// TIA Portal project "Pozycjoner_v7" (V15.1) (continued)
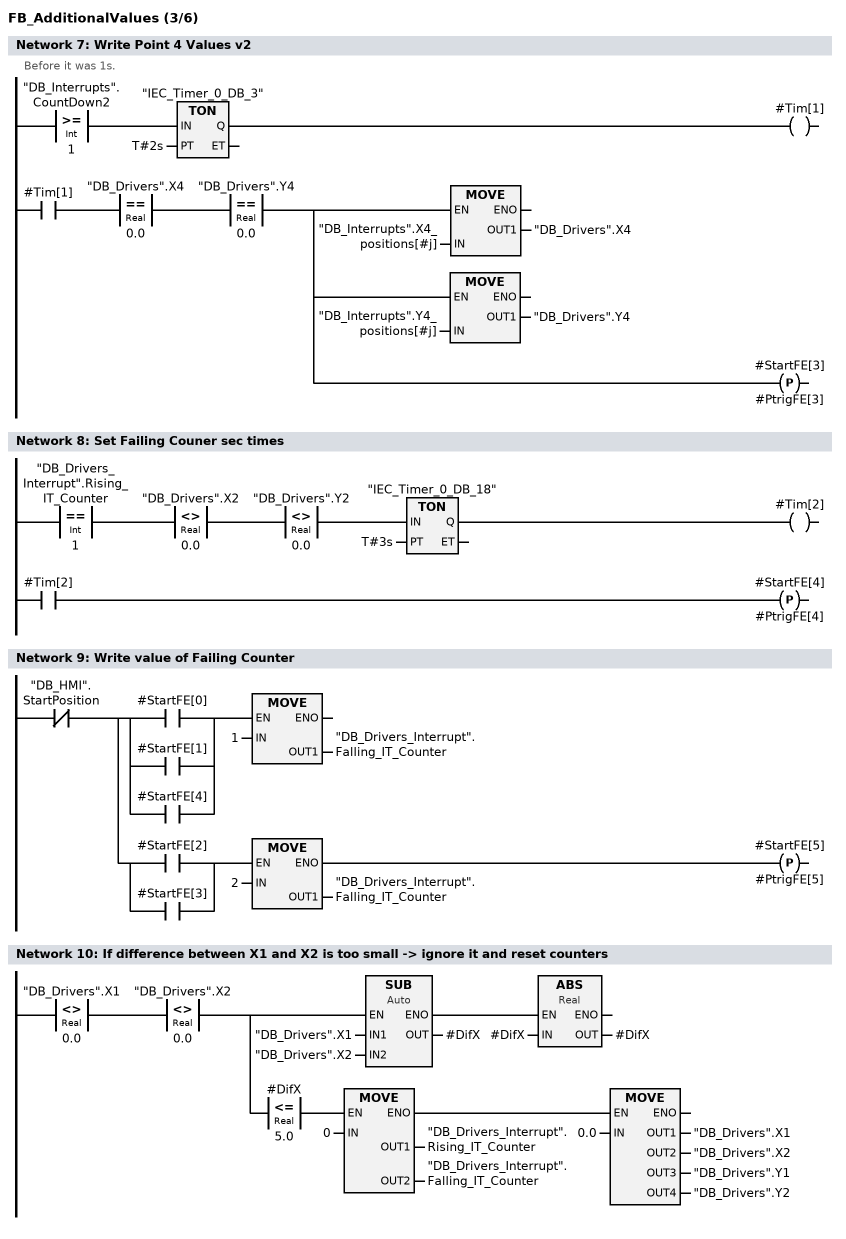
   "IEC_Timer_0_DB_3".TON(IN := "DB_Interrupts".CountDown2 >= 1, PT := T#2s);
   #Tim[1] := "IEC_Timer_0_DB_3".Q;
   #_w1 := #Tim[1] AND ("DB_Drivers".X4 = 0.0) AND ("DB_Drivers".Y4 = 0.0);
   IF #_w1 THEN
       "DB_Drivers".X4 := "DB_Interrupts".X4_positions[#j];
       "DB_Drivers".Y4 := "DB_Interrupts".Y4_positions[#j];
   END_IF;
   #StartFE[3] := #_w1 AND NOT #PtrigFE[3];   // rising edge
   #PtrigFE[3] := #_w1;
END_REGION

REGION Network 8: Set Failing Couner sec times
   "IEC_Timer_0_DB_18".TON(IN := ("DB_Drivers_Interrupt".Rising_IT_Counter = 1) AND ("DB_Drivers".X2 <> 0.0) AND ("DB_Drivers".Y2 <> 0.0),
                           PT := T#3s);
   #Tim[2] := "IEC_Timer_0_DB_18".Q;
   #StartFE[4] := #Tim[2] AND NOT #PtrigFE[4];   // rising edge
   #PtrigFE[4] := #Tim[2];
END_REGION

REGION Network 9: Write value of Failing Counter
   #_w1 := NOT "DB_HMI".StartPosition;
   IF #_w1 AND (#StartFE[0] OR #StartFE[1] OR #StartFE[4]) THEN
       "DB_Drivers_Interrupt".Falling_IT_Counter := 1;
   END_IF;
   #_w2 := #_w1 AND (#StartFE[2] OR #StartFE[3]);
   IF #_w2 THEN "DB_Drivers_Interrupt".Falling_IT_Counter := 2; END_IF;
   #StartFE[5] := #_w2 AND NOT #PtrigFE[5];   // rising edge
   #PtrigFE[5] := #_w2;
END_REGION

REGION Network 10: If difference between X1 and X2 is too small -> ignore it and reset counters
   RUNG wire#powerrail
      { S7_Templates := "SrcType := Real" } NE_Contact(in1 := "DB_Drivers".X1, in2 := 0.0)
      { S7_Templates := "SrcType := Real" } NE_Contact(in1 := "DB_Drivers".X2, in2 := 0.0)
      wire#w1
      Sub(in1 := "DB_Drivers".X1, in2 := "DB_Drivers".X2, out => #DifX)
      { S7_Templates := "SrcType := Real" } Abs(in := #DifX, out => #DifX)
   END_RUNG
   RUNG wire#w1
      { S7_Templates := "SrcType := Real" } LE_Contact(in1 := #DifX, in2 := 5.0)
      Move(in := 0, out1 => "DB_Drivers_Interrupt".Rising_IT_Counter, out2 => "DB_Drivers_Interrupt".Falling_IT_Counter)
      Move(in := 0.0, out1 => "DB_Drivers".X1, out2 => "DB_Drivers".X2, out3 => "DB_Drivers".Y1, out4 => "DB_Drivers".Y2)
   END_RUNG
   // the same network as SCL:
   #_w1 := ("DB_Drivers".X1 <> 0.0) AND ("DB_Drivers".X2 <> 0.0);
   IF #_w1 THEN
       #DifX := "DB_Drivers".X1 - "DB_Drivers".X2;
       #DifX := ABS(#DifX);
   END_IF;
   IF #_w1 AND (#DifX <= 5.0) THEN
       "DB_Drivers_Interrupt".Rising_IT_Counter := 0;
       "DB_Drivers_Interrupt".Falling_IT_Counter := 0;
       "DB_Drivers".X1 := 0.0;
       "DB_Drivers".X2 := 0.0;
       "DB_Drivers".Y1 := 0.0;
       "DB_Drivers".Y2 := 0.0;
   END_IF;
END_REGION

REGION Network 11: Repeat move if rising edge was detected but falling edge counter = 0 for 10 sec
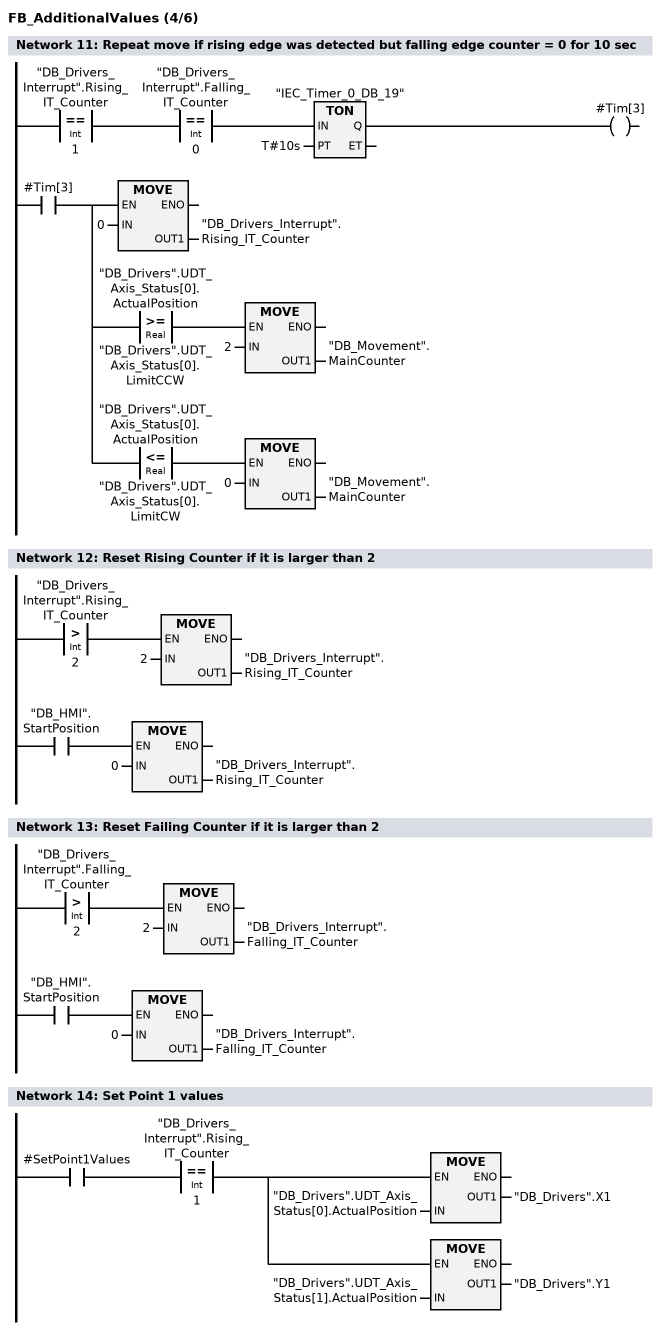
   "IEC_Timer_0_DB_19".TON(IN := ("DB_Drivers_Interrupt".Rising_IT_Counter = 1) AND ("DB_Drivers_Interrupt".Falling_IT_Counter = 0),
                           PT := T#10s);
   #Tim[3] := "IEC_Timer_0_DB_19".Q;
   IF #Tim[3] THEN "DB_Drivers_Interrupt".Rising_IT_Counter := 0; END_IF;
   IF #Tim[3] AND ("DB_Drivers".UDT_Axis_Status[0].ActualPosition >= "DB_Drivers".UDT_Axis_Status[0].LimitCCW) THEN
       "DB_Movement".MainCounter := 2;
   END_IF;
   IF #Tim[3] AND ("DB_Drivers".UDT_Axis_Status[0].ActualPosition <= "DB_Drivers".UDT_Axis_Status[0].LimitCW) THEN
       "DB_Movement".MainCounter := 0;
   END_IF;
END_REGION

REGION Network 12: Reset Rising Counter if it is larger than 2
   RUNG wire#powerrail
      { S7_Templates := "SrcType := Int" } GT_Contact(in1 := "DB_Drivers_Interrupt".Rising_IT_Counter, in2 := 2)
      Move(in := 2, out1 => "DB_Drivers_Interrupt".Rising_IT_Counter)
   END_RUNG
   RUNG wire#powerrail
      Contact( "DB_HMI".StartPosition )
      Move(in := 0, out1 => "DB_Drivers_Interrupt".Rising_IT_Counter)
   END_RUNG
   // the same network as SCL:
   IF "DB_Drivers_Interrupt".Rising_IT_Counter > 2 THEN
       "DB_Drivers_Interrupt".Rising_IT_Counter := 2;
   END_IF;
   IF "DB_HMI".StartPosition THEN "DB_Drivers_Interrupt".Rising_IT_Counter := 0; END_IF;
END_REGION

REGION Network 13: Reset Failing Counter if it is larger than 2
   RUNG wire#powerrail
      { S7_Templates := "SrcType := Int" } GT_Contact(in1 := "DB_Drivers_Interrupt".Falling_IT_Counter, in2 := 2)
      Move(in := 2, out1 => "DB_Drivers_Interrupt".Falling_IT_Counter)
   END_RUNG
   RUNG wire#powerrail
      Contact( "DB_HMI".StartPosition )
      Move(in := 0, out1 => "DB_Drivers_Interrupt".Falling_IT_Counter)
   END_RUNG
   // the same network as SCL:
   IF "DB_Drivers_Interrupt".Falling_IT_Counter > 2 THEN
       "DB_Drivers_Interrupt".Falling_IT_Counter := 2;
   END_IF;
   IF "DB_HMI".StartPosition THEN "DB_Drivers_Interrupt".Falling_IT_Counter := 0; END_IF;
END_REGION

REGION Network 14: Set Point 1 values
   RUNG wire#powerrail
      Contact( #SetPoint1Values )
      { S7_Templates := "SrcType := Int" } EQ_Contact(in1 := "DB_Drivers_Interrupt".Rising_IT_Counter, in2 := 1)
      wire#w1
      Move(in := "DB_Drivers".UDT_Axis_Status[0].ActualPosition, out1 => "DB_Drivers".X1)
   END_RUNG
   RUNG wire#w1
      Move(in := "DB_Drivers".UDT_Axis_Status[1].ActualPosition, out1 => "DB_Drivers".Y1)
   END_RUNG
   // the same network as SCL:
   IF #SetPoint1Values AND ("DB_Drivers_Interrupt".Rising_IT_Counter = 1) THEN
       "DB_Drivers".X1 := "DB_Drivers".UDT_Axis_Status[0].ActualPosition;
       "DB_Drivers".Y1 := "DB_Drivers".UDT_Axis_Status[1].ActualPosition;
   END_IF;
END_REGION

REGION Network 15: Set Point 3 values
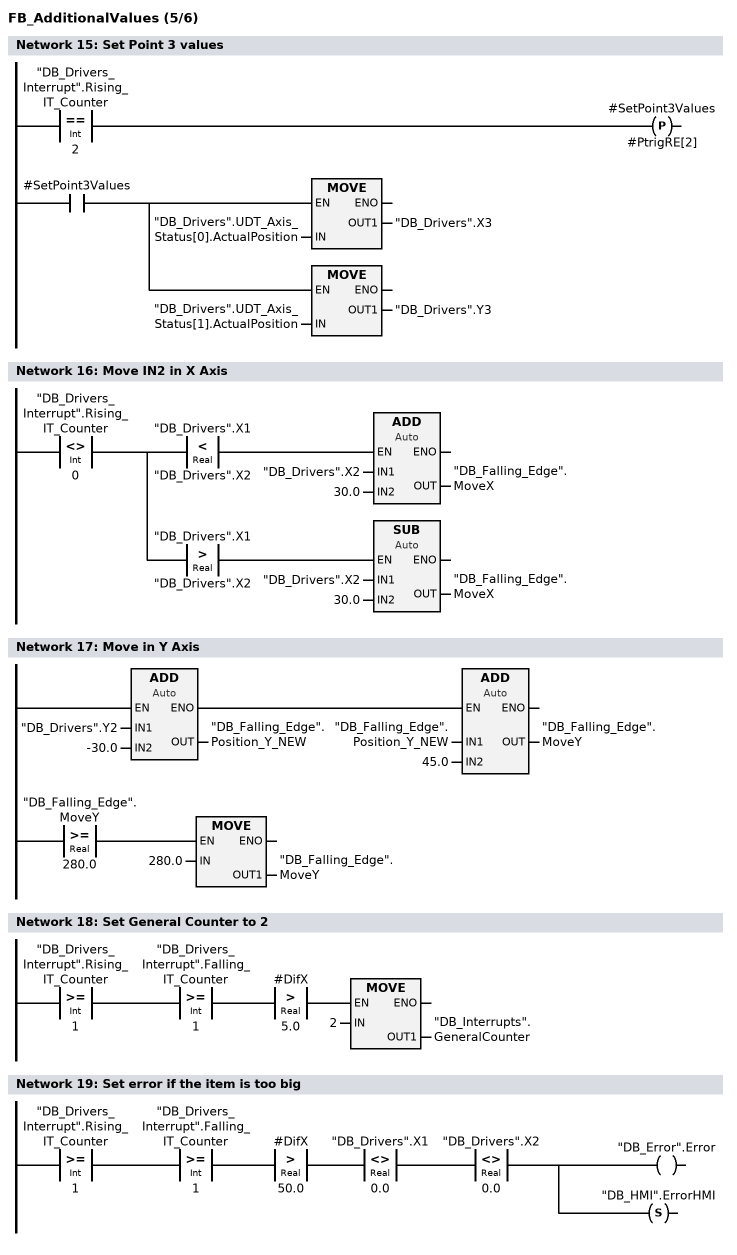
   #_w1 := "DB_Drivers_Interrupt".Rising_IT_Counter = 2;
   #SetPoint3Values := #_w1 AND NOT #PtrigRE[2];   // rising edge
   #PtrigRE[2] := #_w1;
   IF #SetPoint3Values THEN
       "DB_Drivers".X3 := "DB_Drivers".UDT_Axis_Status[0].ActualPosition;
       "DB_Drivers".Y3 := "DB_Drivers".UDT_Axis_Status[1].ActualPosition;
   END_IF;
END_REGION

REGION Network 16: Move IN2 in X Axis
   RUNG wire#powerrail
      { S7_Templates := "SrcType := Int" } NE_Contact(in1 := "DB_Drivers_Interrupt".Rising_IT_Counter, in2 := 0)
      wire#w1
      { S7_Templates := "SrcType := Real" } LT_Contact(in1 := "DB_Drivers".X1, in2 := "DB_Drivers".X2)
      Add(in1 := "DB_Drivers".X2, in2 := 30.0, out => "DB_Falling_Edge".MoveX)
   END_RUNG
   RUNG wire#w1
      { S7_Templates := "SrcType := Real" } GT_Contact(in1 := "DB_Drivers".X1, in2 := "DB_Drivers".X2)
      Sub(in1 := "DB_Drivers".X2, in2 := 30.0, out => "DB_Falling_Edge".MoveX)
   END_RUNG
   // the same network as SCL:
   #_w1 := "DB_Drivers_Interrupt".Rising_IT_Counter <> 0;
   IF #_w1 AND ("DB_Drivers".X1 < "DB_Drivers".X2) THEN
       "DB_Falling_Edge".MoveX := "DB_Drivers".X2 + 30.0;
   END_IF;
   IF #_w1 AND ("DB_Drivers".X1 > "DB_Drivers".X2) THEN
       "DB_Falling_Edge".MoveX := "DB_Drivers".X2 - 30.0;
   END_IF;
END_REGION

REGION Network 17: Move in Y Axis
   RUNG wire#powerrail
      Add(in1 := "DB_Drivers".Y2, in2 := -30.0, out => "DB_Falling_Edge".Position_Y_NEW)
      Add(in1 := "DB_Falling_Edge".Position_Y_NEW, in2 := 45.0, out => "DB_Falling_Edge".MoveY)
   END_RUNG
   RUNG wire#powerrail
      { S7_Templates := "SrcType := Real" } GE_Contact(in1 := "DB_Falling_Edge".MoveY, in2 := 280.0)
      Move(in := 280.0, out1 => "DB_Falling_Edge".MoveY)
   END_RUNG
   // the same network as SCL:
   "DB_Falling_Edge".Position_Y_NEW := "DB_Drivers".Y2 + (-30.0);
   "DB_Falling_Edge".MoveY := "DB_Falling_Edge".Position_Y_NEW + 45.0;
   IF "DB_Falling_Edge".MoveY >= 280.0 THEN "DB_Falling_Edge".MoveY := 280.0; END_IF;
END_REGION

REGION Network 18: Set General Counter to 2
   RUNG wire#powerrail
      { S7_Templates := "SrcType := Int" } GE_Contact(in1 := "DB_Drivers_Interrupt".Rising_IT_Counter, in2 := 1)
      { S7_Templates := "SrcType := Int" } GE_Contact(in1 := "DB_Drivers_Interrupt".Falling_IT_Counter, in2 := 1)
      { S7_Templates := "SrcType := Real" } GT_Contact(in1 := #DifX, in2 := 5.0)
      Move(in := 2, out1 => "DB_Interrupts".GeneralCounter)
   END_RUNG
   // the same network as SCL:
   IF ("DB_Drivers_Interrupt".Rising_IT_Counter >= 1) AND ("DB_Drivers_Interrupt".Falling_IT_Counter >= 1) AND (#DifX > 5.0) THEN
       "DB_Interrupts".GeneralCounter := 2;
   END_IF;
END_REGION

REGION Network 19: Set error if the item is too big
   RUNG wire#powerrail
      { S7_Templates := "SrcType := Int" } GE_Contact(in1 := "DB_Drivers_Interrupt".Rising_IT_Counter, in2 := 1)
      { S7_Templates := "SrcType := Int" } GE_Contact(in1 := "DB_Drivers_Interrupt".Falling_IT_Counter, in2 := 1)
      { S7_Templates := "SrcType := Real" } GT_Contact(in1 := #DifX, in2 := 50.0)
      { S7_Templates := "SrcType := Real" } NE_Contact(in1 := "DB_Drivers".X1, in2 := 0.0)
      { S7_Templates := "SrcType := Real" } NE_Contact(in1 := "DB_Drivers".X2, in2 := 0.0)
      wire#w1
      Coil( "DB_Error".Error )
   END_RUNG
   RUNG wire#w1
      S_Coil( "DB_HMI".ErrorHMI )
   END_RUNG
   // the same network as SCL:
   "DB_Error".Error := ("DB_Drivers_Interrupt".Rising_IT_Counter >= 1) AND ("DB_Drivers_Interrupt".Falling_IT_Counter >= 1) AND (#DifX > 50.0) AND ("DB_Drivers".X1 <> 0.0) AND ("DB_Drivers".X2 <> 0.0);
   IF "DB_Error".Error THEN "DB_HMI".ErrorHMI := TRUE; END_IF;
END_REGION

REGION Network 20: Check the last point once again
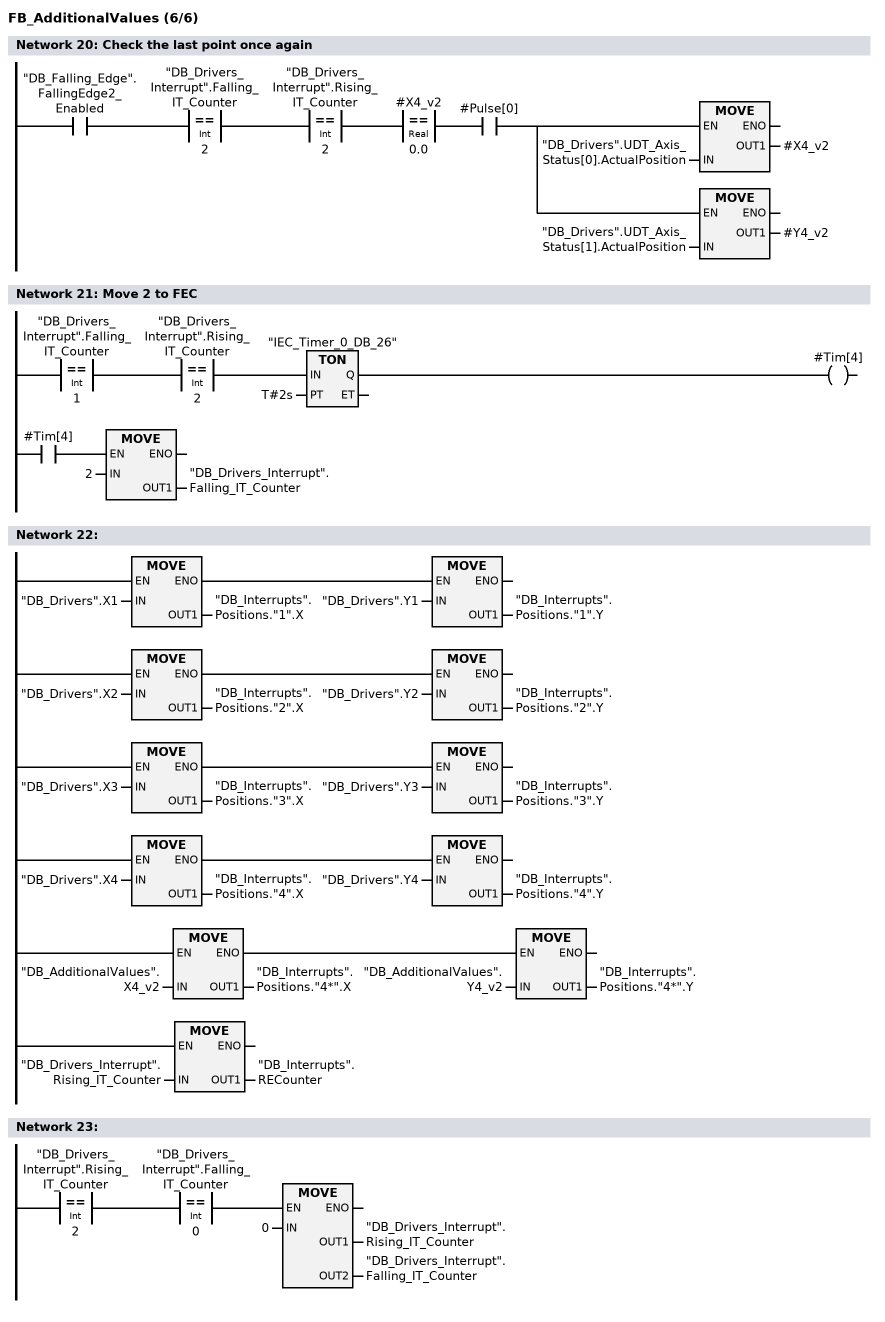
   RUNG wire#powerrail
      Contact( "DB_Falling_Edge".FallingEdge2_Enabled )
      { S7_Templates := "SrcType := Int" } EQ_Contact(in1 := "DB_Drivers_Interrupt".Falling_IT_Counter, in2 := 2)
      { S7_Templates := "SrcType := Int" } EQ_Contact(in1 := "DB_Drivers_Interrupt".Rising_IT_Counter, in2 := 2)
      { S7_Templates := "SrcType := Real" } EQ_Contact(in1 := #X4_v2, in2 := 0.0)
      Contact( #Pulse[0] )
      wire#w1
      Move(in := "DB_Drivers".UDT_Axis_Status[0].ActualPosition, out1 => #X4_v2)
   END_RUNG
   RUNG wire#w1
      Move(in := "DB_Drivers".UDT_Axis_Status[1].ActualPosition, out1 => #Y4_v2)
   END_RUNG
   // the same network as SCL:
   #_w1 := "DB_Falling_Edge".FallingEdge2_Enabled AND ("DB_Drivers_Interrupt".Falling_IT_Counter = 2) AND ("DB_Drivers_Interrupt".Rising_IT_Counter = 2) AND (#X4_v2 = 0.0) AND #Pulse[0];
   IF #_w1 THEN
       #X4_v2 := "DB_Drivers".UDT_Axis_Status[0].ActualPosition;
       #Y4_v2 := "DB_Drivers".UDT_Axis_Status[1].ActualPosition;
   END_IF;
END_REGION

REGION Network 21: Move 2 to FEC
   "IEC_Timer_0_DB_26".TON(IN := ("DB_Drivers_Interrupt".Falling_IT_Counter = 1) AND ("DB_Drivers_Interrupt".Rising_IT_Counter = 2),
                           PT := T#2s);
   #Tim[4] := "IEC_Timer_0_DB_26".Q;
   IF #Tim[4] THEN "DB_Drivers_Interrupt".Falling_IT_Counter := 2; END_IF;
END_REGION

REGION Network 22
   RUNG wire#powerrail
      Move(in := "DB_Drivers".X1, out1 => "DB_Interrupts".Positions."1".X)
      Move(in := "DB_Drivers".Y1, out1 => "DB_Interrupts".Positions."1".Y)
   END_RUNG
   RUNG wire#powerrail
      Move(in := "DB_Drivers".X2, out1 => "DB_Interrupts".Positions."2".X)
      Move(in := "DB_Drivers".Y2, out1 => "DB_Interrupts".Positions."2".Y)
   END_RUNG
   RUNG wire#powerrail
      Move(in := "DB_Drivers".X3, out1 => "DB_Interrupts".Positions."3".X)
      Move(in := "DB_Drivers".Y3, out1 => "DB_Interrupts".Positions."3".Y)
   END_RUNG
   RUNG wire#powerrail
      Move(in := "DB_Drivers".X4, out1 => "DB_Interrupts".Positions."4".X)
      Move(in := "DB_Drivers".Y4, out1 => "DB_Interrupts".Positions."4".Y)
   END_RUNG
   RUNG wire#powerrail
      Move(in := "DB_AdditionalValues".X4_v2, out1 => "DB_Interrupts".Positions."4*".X)
      Move(in := "DB_AdditionalValues".Y4_v2, out1 => "DB_Interrupts".Positions."4*".Y)
   END_RUNG
   RUNG wire#powerrail
      Move(in := "DB_Drivers_Interrupt".Rising_IT_Counter, out1 => "DB_Interrupts".RECounter)
   END_RUNG
   // the same network as SCL:
   "DB_Interrupts".Positions."1".X := "DB_Drivers".X1;
   "DB_Interrupts".Positions."1".Y := "DB_Drivers".Y1;
   "DB_Interrupts".Positions."2".X := "DB_Drivers".X2;
   "DB_Interrupts".Positions."2".Y := "DB_Drivers".Y2;
   "DB_Interrupts".Positions."3".X := "DB_Drivers".X3;
   "DB_Interrupts".Positions."3".Y := "DB_Drivers".Y3;
   "DB_Interrupts".Positions."4".X := "DB_Drivers".X4;
   "DB_Interrupts".Positions."4".Y := "DB_Drivers".Y4;
   "DB_Interrupts".Positions."4*".X := "DB_AdditionalValues".X4_v2;
   "DB_Interrupts".Positions."4*".Y := "DB_AdditionalValues".Y4_v2;
   "DB_Interrupts".RECounter := "DB_Drivers_Interrupt".Rising_IT_Counter;
END_REGION

REGION Network 23
   RUNG wire#powerrail
      { S7_Templates := "SrcType := Int" } EQ_Contact(in1 := "DB_Drivers_Interrupt".Rising_IT_Counter, in2 := 2)
      { S7_Templates := "SrcType := Int" } EQ_Contact(in1 := "DB_Drivers_Interrupt".Falling_IT_Counter, in2 := 0)
      Move(in := 0, out1 => "DB_Drivers_Interrupt".Rising_IT_Counter, out2 => "DB_Drivers_Interrupt".Falling_IT_Counter)
   END_RUNG
   // the same network as SCL:
   IF ("DB_Drivers_Interrupt".Rising_IT_Counter = 2) AND ("DB_Drivers_Interrupt".Falling_IT_Counter = 0) THEN
       "DB_Drivers_Interrupt".Rising_IT_Counter := 0;
       "DB_Drivers_Interrupt".Falling_IT_Counter := 0;
   END_IF;
END_REGION
END_FUNCTION_BLOCK

FUNCTION_BLOCK "FB_Falling_Edge"   // FB9, LAD
{ S7_Optimized_Access := 'TRUE' }
VERSION : 0.1
   VAR_INPUT
      LaserSensor : Bool;
   END_VAR
   VAR
      X_Position2 : Real;
      Y_Position2 : Real;
      Position_Y_NEW : Real;   // New Y position
      MoveX : Real;   // Keep moving after detecting item
      UDT_AxisControl : Array[0..2] of "UDT_AxisControl";
      UDT_AxisStatus : Array[0..2] of "UDT_AxisStatus";
      Y_MIN : Int;
      Y_MAX : Real;
      MoveX_MIN : Int;
      MoveX_MAX : Int;
      MoveY : Real;
      MainCounter : Int;
      Enabled : Bool;
      moveY_min : Int;
      moveY_max : Int;
      FallingEdge2_Enabled : Bool;
      StartX : Array[0..2] of Bool;
      StartY : Array[0..2] of Bool;
      PtrigX : Array[0..2] of Bool;
      PtrigY : Array[0..2] of Bool;
      Timers : Array[0..2] of Bool;
   END_VAR
   VAR_TEMP   // added for the SCL form of the ladder/FBD networks
      _w1 : Bool;
   END_VAR
BEGIN

REGION Network 1: Enabled
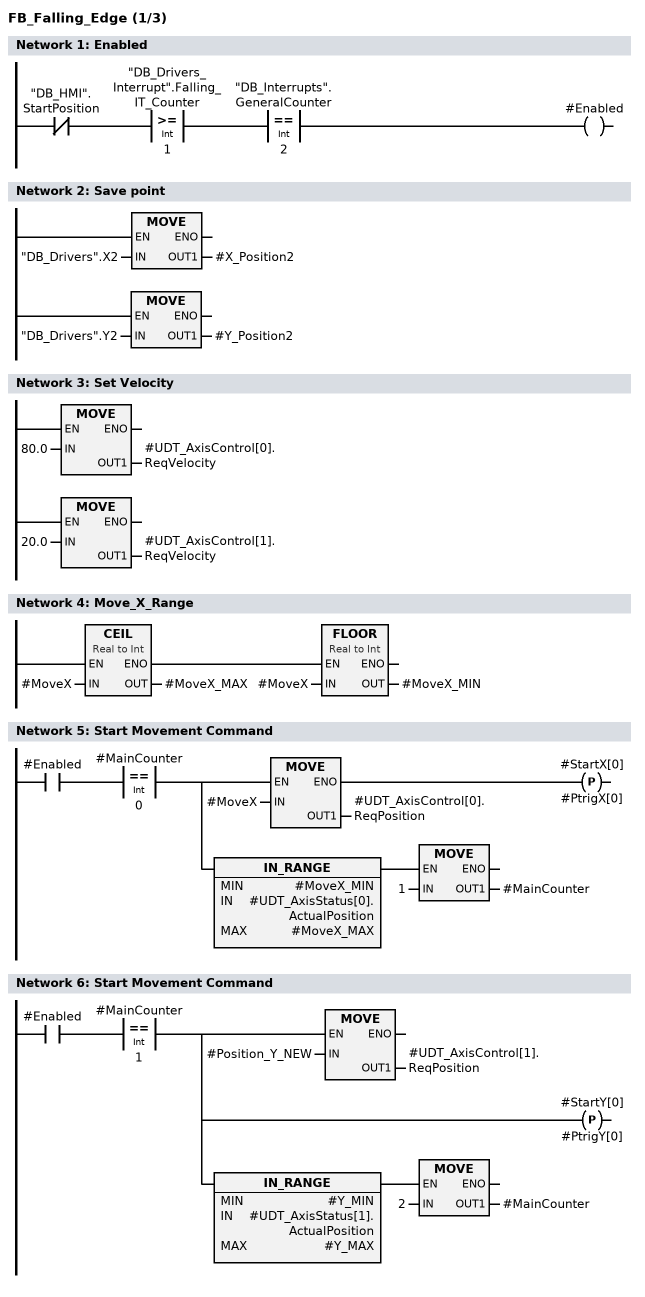
   RUNG wire#powerrail
      I_Contact( "DB_HMI".StartPosition )
      { S7_Templates := "SrcType := Int" } GE_Contact(in1 := "DB_Drivers_Interrupt".Falling_IT_Counter, in2 := 1)
      { S7_Templates := "SrcType := Int" } EQ_Contact(in1 := "DB_Interrupts".GeneralCounter, in2 := 2)
      Coil( #Enabled )
   END_RUNG
   // the same network as SCL:
   #Enabled := NOT "DB_HMI".StartPosition AND ("DB_Drivers_Interrupt".Falling_IT_Counter >= 1) AND ("DB_Interrupts".GeneralCounter = 2);
END_REGION

REGION Network 2: Save point
   RUNG wire#powerrail
      Move(in := "DB_Drivers".X2, out1 => #X_Position2)
   END_RUNG
   RUNG wire#powerrail
      Move(in := "DB_Drivers".Y2, out1 => #Y_Position2)
   END_RUNG
   // the same network as SCL:
   #X_Position2 := "DB_Drivers".X2;
   #Y_Position2 := "DB_Drivers".Y2;
END_REGION

REGION Network 3: Set Velocity
   RUNG wire#powerrail
      Move(in := 80.0, out1 => #UDT_AxisControl[0].ReqVelocity)
   END_RUNG
   RUNG wire#powerrail
      Move(in := 20.0, out1 => #UDT_AxisControl[1].ReqVelocity)
   END_RUNG
   // the same network as SCL:
   #UDT_AxisControl[0].ReqVelocity := 80.0;
   #UDT_AxisControl[1].ReqVelocity := 20.0;
END_REGION

REGION Network 4: Move_X_Range
   #MoveX_MAX := CEIL(#MoveX);
   #MoveX_MIN := FLOOR(#MoveX);
END_REGION

REGION Network 5: Start Movement Command
   #_w1 := #Enabled AND (#MainCounter = 0);
   IF #_w1 THEN #UDT_AxisControl[0].ReqPosition := #MoveX; END_IF;
   #StartX[0] := #_w1 AND NOT #PtrigX[0];   // rising edge
   #PtrigX[0] := #_w1;
   IF #_w1 AND (#MoveX_MIN <= #UDT_AxisStatus[0].ActualPosition) AND (#UDT_AxisStatus[0].ActualPosition <= #MoveX_MAX) THEN
       #MainCounter := 1;
   END_IF;
END_REGION

REGION Network 6: Start Movement Command
   #_w1 := #Enabled AND (#MainCounter = 1);
   IF #_w1 THEN #UDT_AxisControl[1].ReqPosition := #Position_Y_NEW; END_IF;
   #StartY[0] := #_w1 AND NOT #PtrigY[0];   // rising edge
   #PtrigY[0] := #_w1;
   IF #_w1 AND (#Y_MIN <= #UDT_AxisStatus[1].ActualPosition) AND (#UDT_AxisStatus[1].ActualPosition <= #Y_MAX) THEN
       #MainCounter := 2;
   END_IF;
END_REGION

REGION Network 7: NewPositionY Range
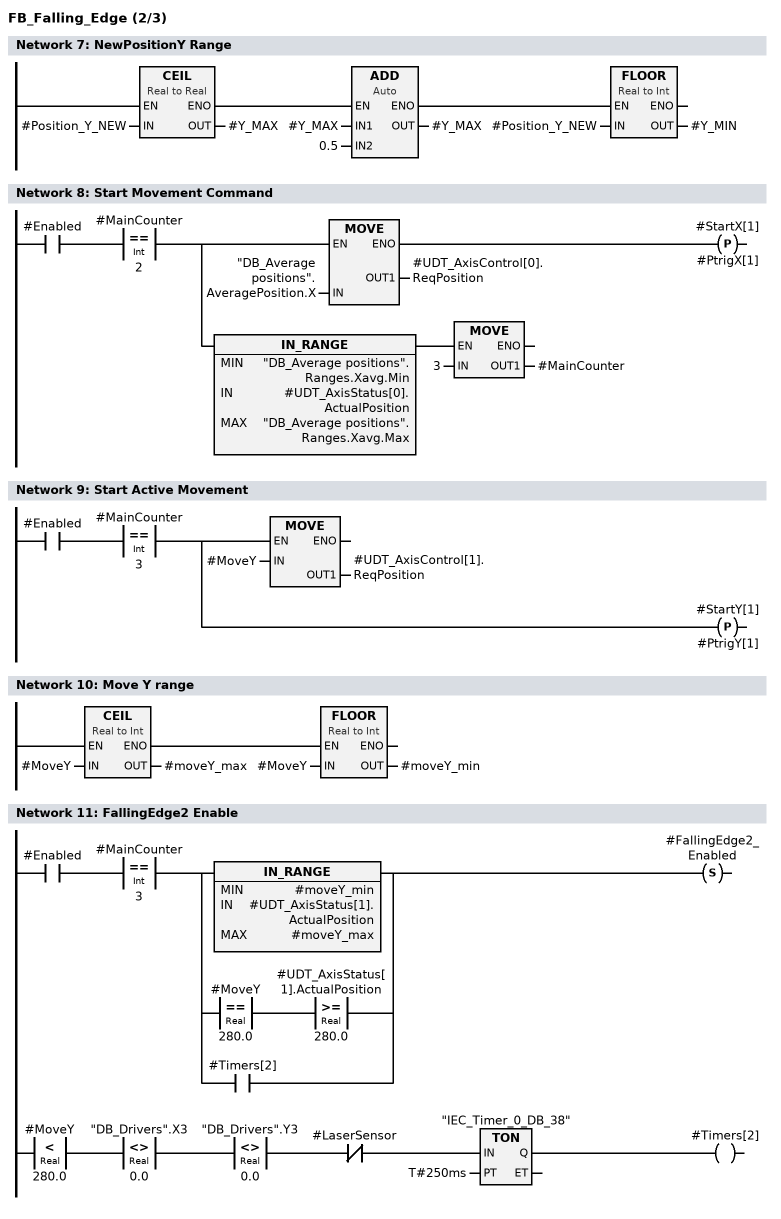
   #Y_MAX := CEIL(#Position_Y_NEW);
   #Y_MAX := #Y_MAX + 0.5;
   #Y_MIN := FLOOR(#Position_Y_NEW);
END_REGION

REGION Network 8: Start Movement Command
   #_w1 := #Enabled AND (#MainCounter = 2);
   IF #_w1 THEN #UDT_AxisControl[0].ReqPosition := "DB_Average positions".AveragePosition.X; END_IF;
   #StartX[1] := #_w1 AND NOT #PtrigX[1];   // rising edge
   #PtrigX[1] := #_w1;
   IF #_w1 AND ("DB_Average positions".Ranges.Xavg.Min <= #UDT_AxisStatus[0].ActualPosition) AND (#UDT_AxisStatus[0].ActualPosition <= "DB_Average positions".Ranges.Xavg.Max) THEN
       #MainCounter := 3;
   END_IF;
END_REGION

REGION Network 9: Start Active Movement
   #_w1 := #Enabled AND (#MainCounter = 3);
   IF #_w1 THEN #UDT_AxisControl[1].ReqPosition := #MoveY; END_IF;
   #StartY[1] := #_w1 AND NOT #PtrigY[1];   // rising edge
   #PtrigY[1] := #_w1;
END_REGION

REGION Network 10: Move Y range
   #moveY_max := CEIL(#MoveY);
   #moveY_min := FLOOR(#MoveY);
END_REGION

REGION Network 11: FallingEdge2 Enable
   IF #Enabled AND (#MainCounter = 3) AND (((#moveY_min <= #UDT_AxisStatus[1].ActualPosition) AND (#UDT_AxisStatus[1].ActualPosition <= #moveY_max)) OR ((#MoveY = 280.0) AND (#UDT_AxisStatus[1].ActualPosition >= 280.0)) OR #Timers[2]) THEN
       #FallingEdge2_Enabled := TRUE;
   END_IF;
   "IEC_Timer_0_DB_38".TON(IN := (#MoveY < 280.0) AND ("DB_Drivers".X3 <> 0.0) AND ("DB_Drivers".Y3 <> 0.0) AND NOT #LaserSensor,
                           PT := T#250ms);
   #Timers[2] := "IEC_Timer_0_DB_38".Q;
END_REGION

REGION Network 12: Start Movement Command
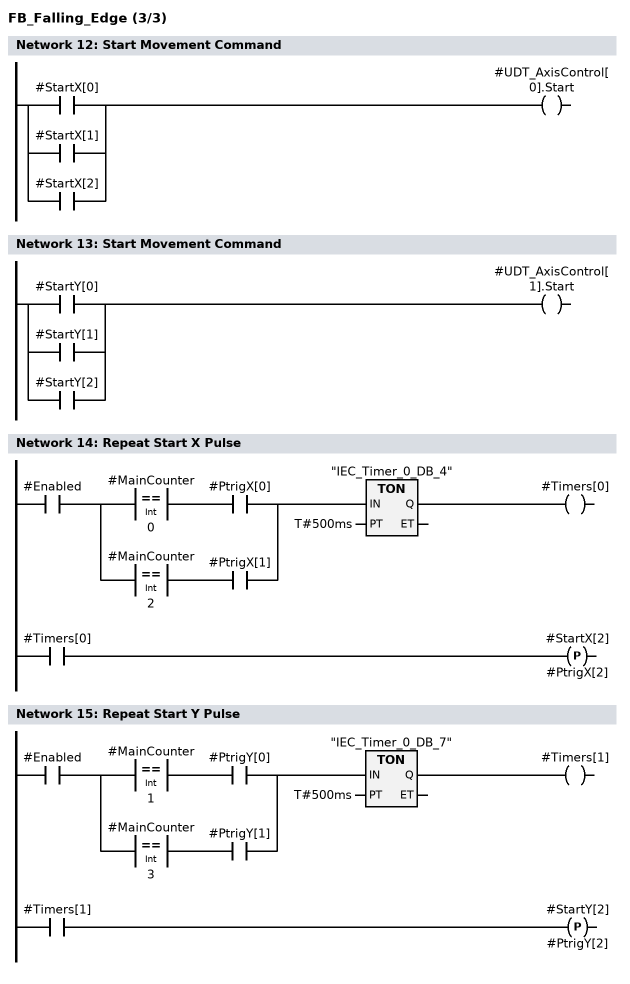
   RUNG wire#powerrail
      Contact( #StartX[0] )
      wire#w1
      Coil( #UDT_AxisControl[0].Start )
   END_RUNG
   RUNG wire#powerrail
      Contact( #StartX[1] )
   END_RUNG wire#w1
   RUNG wire#powerrail
      Contact( #StartX[2] )
   END_RUNG wire#w1
   // the same network as SCL:
   #UDT_AxisControl[0].Start := #StartX[0] OR #StartX[1] OR #StartX[2];
END_REGION

REGION Network 13: Start Movement Command
   RUNG wire#powerrail
      Contact( #StartY[0] )
      wire#w1
      Coil( #UDT_AxisControl[1].Start )
   END_RUNG
   RUNG wire#powerrail
      Contact( #StartY[1] )
   END_RUNG wire#w1
   RUNG wire#powerrail
      Contact( #StartY[2] )
   END_RUNG wire#w1
   // the same network as SCL:
   #UDT_AxisControl[1].Start := #StartY[0] OR #StartY[1] OR #StartY[2];
END_REGION

REGION Network 14: Repeat Start X Pulse
   "IEC_Timer_0_DB_4".TON(IN := #Enabled AND (((#MainCounter = 0) AND #PtrigX[0]) OR ((#MainCounter = 2) AND #PtrigX[1])),
                          PT := T#500ms);
   #Timers[0] := "IEC_Timer_0_DB_4".Q;
   #StartX[2] := #Timers[0] AND NOT #PtrigX[2];   // rising edge
   #PtrigX[2] := #Timers[0];
END_REGION

REGION Network 15: Repeat Start Y Pulse
   "IEC_Timer_0_DB_7".TON(IN := #Enabled AND (((#MainCounter = 1) AND #PtrigY[0]) OR ((#MainCounter = 3) AND #PtrigY[1])),
                          PT := T#500ms);
   #Timers[1] := "IEC_Timer_0_DB_7".Q;
   #StartY[2] := #Timers[1] AND NOT #PtrigY[2];   // rising edge
   #PtrigY[2] := #Timers[1];
END_REGION
END_FUNCTION_BLOCK

// folder: Displacement/Center Point Calculation/Line2

FUNCTION_BLOCK "FB_Line2"   // FB11, LAD
{ S7_Optimized_Access := 'TRUE' }
VERSION : 0.1
   VAR_INPUT
      LaserSensor : Bool;
   END_VAR
   VAR
      UDT_AxisControl : Array[0..2] of "UDT_AxisControl";
      UDT_AxisStatus : Array[0..2] of "UDT_AxisStatus";
      Ranges : Struct
         X_MAX : Real;
         X_MIN : Real;
         Y_MAX : Real;
         Y_MIN : Real;
      END_STRUCT;
      StartX : Array[0..3] of Bool;
      PtrigX : Array[0..3] of Bool;
      StartY : Array[0..4] of Bool;
      PtrigY : Array[0..4] of Bool;
      Enabled : Bool;
      Midpoint : Bool;
      Tim : Array[0..5] of Bool;
   END_VAR
   VAR_TEMP   // added for the SCL form of the ladder/FBD networks
      _w1 : Bool;
      _w2 : Bool;
   END_VAR
BEGIN

REGION Network 1: Enabled block
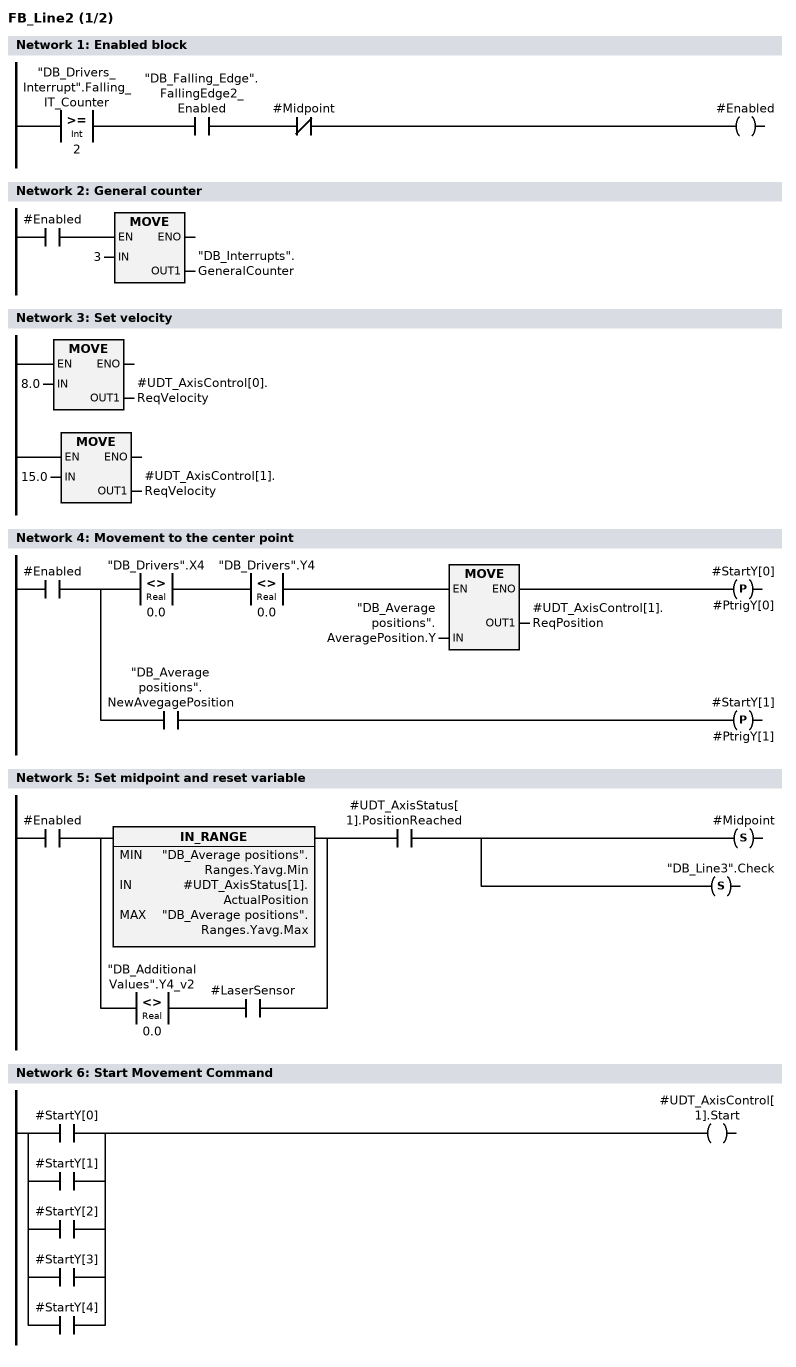
   RUNG wire#powerrail
      { S7_Templates := "SrcType := Int" } GE_Contact(in1 := "DB_Drivers_Interrupt".Falling_IT_Counter, in2 := 2)
      Contact( "DB_Falling_Edge".FallingEdge2_Enabled )
      I_Contact( #Midpoint )
      Coil( #Enabled )
   END_RUNG
   // the same network as SCL:
   #Enabled := ("DB_Drivers_Interrupt".Falling_IT_Counter >= 2) AND "DB_Falling_Edge".FallingEdge2_Enabled AND NOT #Midpoint;
END_REGION

REGION Network 2: General counter
   RUNG wire#powerrail
      Contact( #Enabled )
      Move(in := 3, out1 => "DB_Interrupts".GeneralCounter)
   END_RUNG
   // the same network as SCL:
   IF #Enabled THEN "DB_Interrupts".GeneralCounter := 3; END_IF;
END_REGION

REGION Network 3: Set velocity
   RUNG wire#powerrail
      Move(in := 8.0, out1 => #UDT_AxisControl[0].ReqVelocity)
   END_RUNG
   RUNG wire#powerrail
      Move(in := 15.0, out1 => #UDT_AxisControl[1].ReqVelocity)
   END_RUNG
   // the same network as SCL:
   #UDT_AxisControl[0].ReqVelocity := 8.0;
   #UDT_AxisControl[1].ReqVelocity := 15.0;
END_REGION

REGION Network 4: Movement to the center point
   #_w1 := #Enabled AND ("DB_Drivers".X4 <> 0.0) AND ("DB_Drivers".Y4 <> 0.0);
   IF #_w1 THEN #UDT_AxisControl[1].ReqPosition := "DB_Average positions".AveragePosition.Y; END_IF;
   #StartY[0] := #_w1 AND NOT #PtrigY[0];   // rising edge
   #PtrigY[0] := #_w1;
   #_w2 := #Enabled AND "DB_Average positions".NewAvegagePosition;
   #StartY[1] := #_w2 AND NOT #PtrigY[1];   // rising edge
   #PtrigY[1] := #_w2;
END_REGION

REGION Network 5: Set midpoint and reset variable
   RUNG wire#powerrail
      Contact( #Enabled )
      wire#w1
      { S7_Templates := "SrcType := Real" } InRange(min := "DB_Average positions".Ranges.Yavg.Min, in := #UDT_AxisStatus[1].ActualPosition, max := "DB_Average positions".Ranges.Yavg.Max)
      wire#w2
      Contact( #UDT_AxisStatus[1].PositionReached )
      wire#w3
      S_Coil( #Midpoint )
   END_RUNG
   RUNG wire#w1
      { S7_Templates := "SrcType := Real" } NE_Contact(in1 := "DB_AdditionalValues".Y4_v2, in2 := 0.0)
      Contact( #LaserSensor )
   END_RUNG wire#w2
   RUNG wire#w3
      S_Coil( "DB_Line3".Check )
   END_RUNG
   // the same network as SCL:
   IF #Enabled AND ((("DB_Average positions".Ranges.Yavg.Min <= #UDT_AxisStatus[1].ActualPosition) AND (#UDT_AxisStatus[1].ActualPosition <= "DB_Average positions".Ranges.Yavg.Max)) OR (("DB_AdditionalValues".Y4_v2 <> 0.0) AND #LaserSensor)) AND #UDT_AxisStatus[1].PositionReached THEN
       #Midpoint := TRUE;
       "DB_Line3".Check := TRUE;
   END_IF;
END_REGION

REGION Network 6: Start Movement Command
   RUNG wire#powerrail
      Contact( #StartY[0] )
      wire#w1
      Coil( #UDT_AxisControl[1].Start )
   END_RUNG
   RUNG wire#powerrail
      Contact( #StartY[1] )
   END_RUNG wire#w1
   RUNG wire#powerrail
      Contact( #StartY[2] )
   END_RUNG wire#w1
   RUNG wire#powerrail
      Contact( #StartY[3] )
   END_RUNG wire#w1
   RUNG wire#powerrail
      Contact( #StartY[4] )
   END_RUNG wire#w1
   // the same network as SCL:
   #UDT_AxisControl[1].Start := #StartY[0] OR #StartY[1] OR #StartY[2] OR #StartY[3] OR #StartY[4];
END_REGION

REGION Network 7: Repeat pulse Y Axis
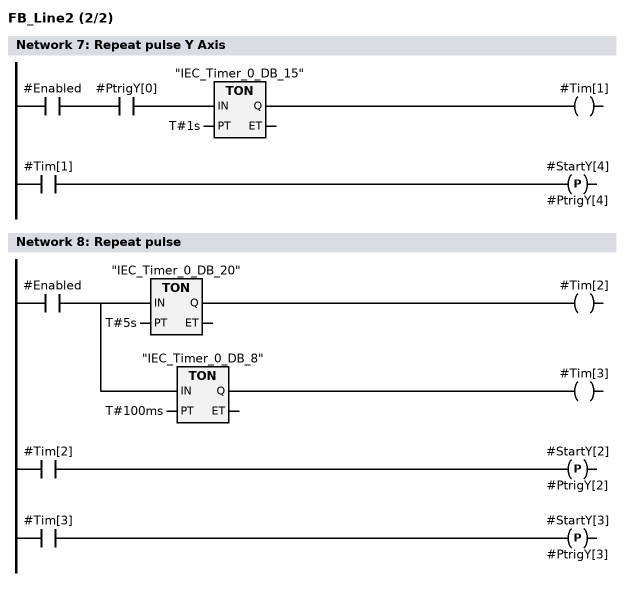
   "IEC_Timer_0_DB_15".TON(IN := #Enabled AND #PtrigY[0], PT := T#1s);
   #Tim[1] := "IEC_Timer_0_DB_15".Q;
   #StartY[4] := #Tim[1] AND NOT #PtrigY[4];   // rising edge
   #PtrigY[4] := #Tim[1];
END_REGION

REGION Network 8: Repeat pulse
   "IEC_Timer_0_DB_20".TON(IN := #Enabled, PT := T#5s);
   #Tim[2] := "IEC_Timer_0_DB_20".Q;
   "IEC_Timer_0_DB_8".TON(IN := #Enabled, PT := T#100ms);
   #Tim[3] := "IEC_Timer_0_DB_8".Q;
   #StartY[2] := #Tim[2] AND NOT #PtrigY[2];   // rising edge
   #PtrigY[2] := #Tim[2];
   #StartY[3] := #Tim[3] AND NOT #PtrigY[3];   // rising edge
   #PtrigY[3] := #Tim[3];
END_REGION
END_FUNCTION_BLOCK

// folder: Displacement/Center Point Calculation/Line3

FUNCTION_BLOCK "FB_Line3"   // FB13, LAD
{ S7_Optimized_Access := 'TRUE' }
VERSION : 0.1
   VAR_INPUT
      LaserSensor : Bool;
   END_VAR
   VAR
      Enabled : Bool;
      MainCounter : Int;
      UDT_AxisCountrol : Array[0..2] of "UDT_AxisControl";
      UDT_AxisStatus : Array[0..2] of "UDT_AxisStatus";
      Line1 : Struct
         X1 : Real;
         Y1 : Real;
         X2 : Real;
         Y2 : Real;
      END_STRUCT;
      Line2 : Struct
         X3 : Real;
         Y3 : Real;
         X4 : Real;
         Y4 : Real;
      END_STRUCT;
      Line3 : Struct
         X5 : Real;
         Y5 : Real;
         X6 : Real;
         Y6 : Real;
      END_STRUCT;
      Check : Bool;
      DiffResult : Real;   // Difference between Yavg and line1
      ShiftDifValue : Real;
      StartX : Array[0..11] of Bool;
      StartY : Array[0..9] of Bool;
      PtrigX : Array[0..11] of Bool;
      PtrigY : Array[0..9] of Bool;
      ShiftDifMin : Real;
      ShiftDifMax : Real;
      MoveXRight : Real;
      MoveXLeft : Real;
      Stop : Array[0..3] of Bool;
      Ntrig : Array[0..1] of Bool;
      Ptrig : Array[0..1] of Bool;
      XavgLine3 : Real;
      GeneralXavg : Real;
      MoveToCenterPoint : Bool;
      YavgRanges : Struct
         Min : Real;
         Max : Real;
      END_STRUCT;
      XavgRanges : Struct
         Min : Real;
         Max : Real;
      END_STRUCT;
      DisplEnabled : Bool;
      Ptrigg : Bool;
      SetCounter : Bool;
      Ptrig1 : Bool;
      SetCount1 : Bool;
      RECountLine3 : Int;
      StartMoveCent : Bool;
      SMCPtrig : Bool;
      MoveToCenter_IR : Bool;
      Midpoint : Bool;
      "Timer" : Bool;
   END_VAR
   VAR_TEMP   // added for the SCL form of the ladder/FBD networks
      _w1 : Bool;
      _w2 : Bool;
   END_VAR
BEGIN

REGION Network 1: Enabled
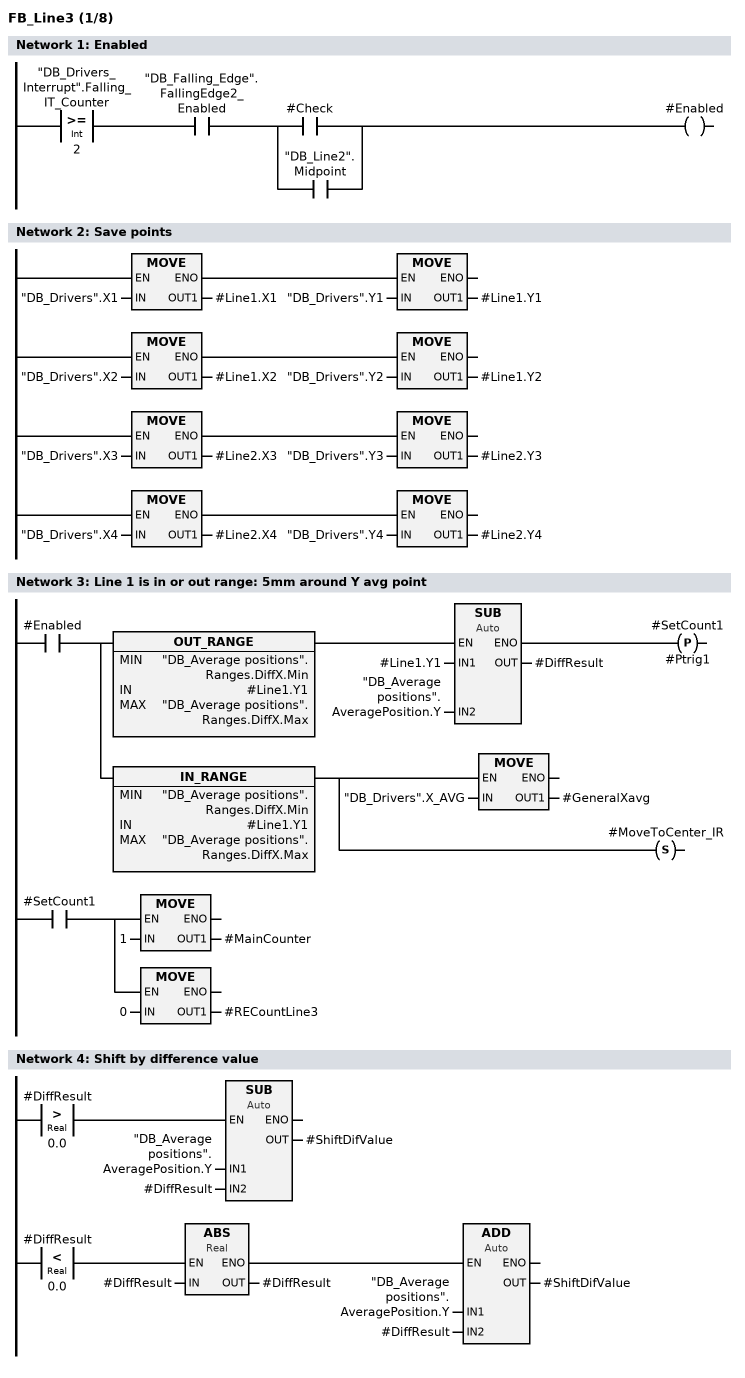
   RUNG wire#powerrail
      { S7_Templates := "SrcType := Int" } GE_Contact(in1 := "DB_Drivers_Interrupt".Falling_IT_Counter, in2 := 2)
      Contact( "DB_Falling_Edge".FallingEdge2_Enabled )
      wire#w1
      Contact( #Check )
      wire#w2
      Coil( #Enabled )
   END_RUNG
   RUNG wire#w1
      Contact( "DB_Line2".Midpoint )
   END_RUNG wire#w2
   // the same network as SCL:
   #Enabled := ("DB_Drivers_Interrupt".Falling_IT_Counter >= 2) AND "DB_Falling_Edge".FallingEdge2_Enabled AND (#Check OR "DB_Line2".Midpoint);
END_REGION

REGION Network 2: Save points
   RUNG wire#powerrail
      Move(in := "DB_Drivers".X1, out1 => #Line1.X1)
      Move(in := "DB_Drivers".Y1, out1 => #Line1.Y1)
   END_RUNG
   RUNG wire#powerrail
      Move(in := "DB_Drivers".X2, out1 => #Line1.X2)
      Move(in := "DB_Drivers".Y2, out1 => #Line1.Y2)
   END_RUNG
   RUNG wire#powerrail
      Move(in := "DB_Drivers".X3, out1 => #Line2.X3)
      Move(in := "DB_Drivers".Y3, out1 => #Line2.Y3)
   END_RUNG
   RUNG wire#powerrail
      Move(in := "DB_Drivers".X4, out1 => #Line2.X4)
      Move(in := "DB_Drivers".Y4, out1 => #Line2.Y4)
   END_RUNG
   // the same network as SCL:
   #Line1.X1 := "DB_Drivers".X1;
   #Line1.Y1 := "DB_Drivers".Y1;
   #Line1.X2 := "DB_Drivers".X2;
   #Line1.Y2 := "DB_Drivers".Y2;
   #Line2.X3 := "DB_Drivers".X3;
   #Line2.Y3 := "DB_Drivers".Y3;
   #Line2.X4 := "DB_Drivers".X4;
   #Line2.Y4 := "DB_Drivers".Y4;
END_REGION
